(* Logix 5000 project; controller PLC_MCC1300_75F1 vendor 1 type 14 code 166 rev 32.11; software revision 32.04; part 27 of 83 *)
(* tags used below, declared in another part *)
   GP_OB_InitializeMain : GP_OB_Initialize;
   M302SpeedUp : MAC_SpeedUp;
   M351 : MAC_Conveyor;
   M352 : MAC_Conveyor;
   M352_ALM : MAC_Conveyor_ALM;
   M352_Data : UDT_Convoy_SL;
   M352_HMR : MAC_Conveyor_HMR;
   M352_HMW : MAC_Conveyor_HMW;
   M352_INPUT_xSLFanOn : BOOL;
   M352_M1_DR : AXIS_CIP_DRIVE;
   M352_M1_DR_IN_MAJ : MOTION_INSTRUCTION;
   M352_M1_DR_IN_MAR : MOTION_INSTRUCTION;
   M352_M1_DR_IN_MAS : MOTION_INSTRUCTION;
   M352_M1_DR_IN_MRP : MOTION_INSTRUCTION;
   M352_M1_DR_MAFR : MOTION_INSTRUCTION;
   M352_M1_DR_MDR : MOTION_INSTRUCTION;
   M352_M1_DR_MSF : MOTION_INSTRUCTION;
   M352_M1_DR_MSO : MOTION_INSTRUCTION;
   M352_M1_DR_OUT_MAJ : MOTION_INSTRUCTION;
   M352_M1_DR_OUT_MAM : MOTION_INSTRUCTION;
   M352_M1_DR_OUT_MAR : MOTION_INSTRUCTION;
   M352_M1_DR_OUT_MAS : MOTION_INSTRUCTION;
   M352_M1_DR_OUT_MCD : MOTION_INSTRUCTION;
   M352_M1_DR_OUT_MRP : MOTION_INSTRUCTION;
   M352_ONS1 : BOOL;
   M352_Output_xAutoMode : BOOL;
   M352_Output_xDescentBlockGlass : BOOL;
   M352_Output_xGlassPresence : BOOL;
   M352_Output_xHA_Alarm : BOOL;   // W254HA1. Acustic alarm
   M352_Output_xHL_Alarm : BOOL;
   M352_Output_xRiseBlockGlass : BOOL;
   M352_SpaceConv_Utilities : SpaceConv_Utilities;
   TMP_d : DINT;
   TMP_dDirection : DINT;
   TMP_r : REAL;
   TMP_rAcc : REAL;
   TMP_rDec : REAL;
   TMP_rSpeed : REAL;
   TMP_rTarget_M1 : REAL;
   TMP_xForwardCommadnForCleaningZone : BOOL;
   TMP_xPositioning : BOOL;
   TMP_xPositioning_M1 : BOOL;
   TMP_xPowerSaving : BOOL;
   TMP_xReverse : BOOL;
   TMP_xReverse_M1 : BOOL;
   TMP_xRun : BOOL;
   TMP_xRun_M1 : BOOL;
   xAlwaysOFF : BOOL;
   Z300_Conveyor : UDT_StandConv[29];
   Z300_Conveyor_Conf : UDT_Conveyor_Config[29];
   Z300_Conveyor_HMW : MAC_Conveyor_ZC_HMW[29];
   Z300_Conveyor_IN_MOTION : MAC_Conveyor_ZC_IN_MOTION[29];
   Z301_HMR : MAC_Zone_ML_HMR;
   Z900 : MAC_Zone;
   Z900_HMW : MAC_Zone_HMW;
(* CommandLogic, continued *)

ROUTINE M352_Output   (* ladder *)
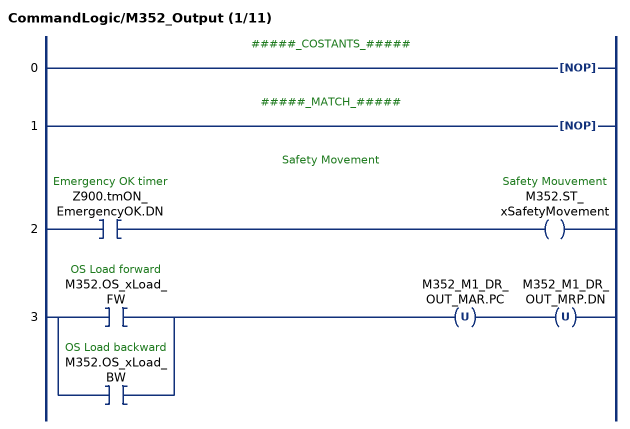
   // #####_COSTANTS_#####
   0: NOP();
   // #####_MATCH_#####
   1: NOP();
   // Safety Movement
   2: XIC(Z900.tmON_EmergencyOK.DN)OTE(M352.ST_xSafetyMovement);
   3: [XIC(M352.OS_xLoad_FW) ,XIC(M352.OS_xLoad_BW) ]OTU(M352_M1_DR_OUT_MAR.PC)OTU(M352_M1_DR_OUT_MRP.DN);
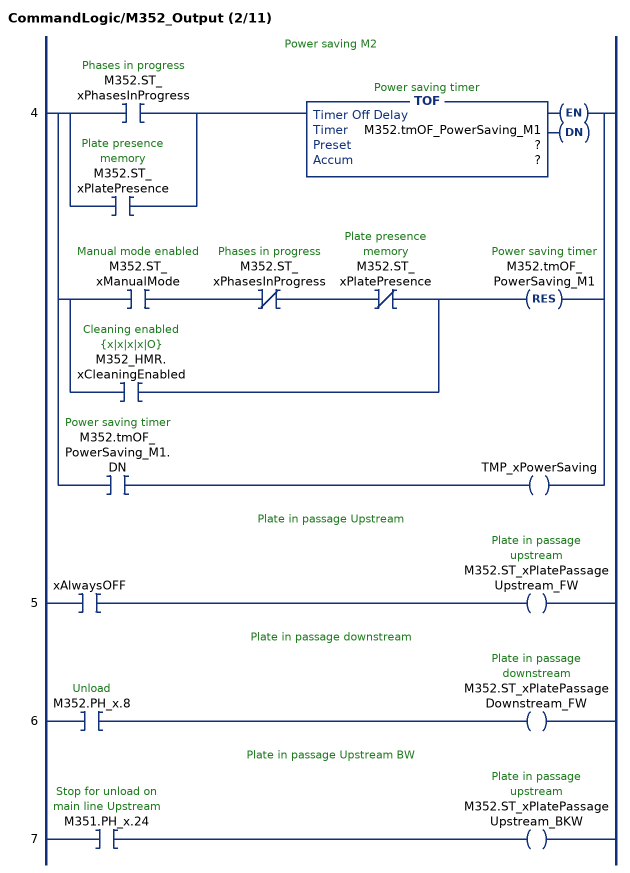
   // Power saving M2
   4: [[XIC(M352.ST_xPhasesInProgress) ,XIC(M352.ST_xPlatePresence) ] TOF(M352.tmOF_PowerSaving_M1,?,?) ,[XIC(M352.ST_xManualMode) XIO(M352.ST_xPhasesInProgress) XIO(M352.ST_xPlatePresence) ,XIC(M352_HMR.xCleaningEnabled) ] RES(M352.tmOF_PowerSaving_M1) ,XIC(M352.tmOF_PowerSaving_M1.DN) OTE(TMP_xPowerSaving) ];
   // Plate in passage Upstream
   5: XIC(xAlwaysOFF)OTE(M352.ST_xPlatePassageUpstream_FW);
   // Plate in passage downstream
   6: XIC(M352.PH_x.8)OTE(M352.ST_xPlatePassageDownstream_FW);
   // Plate in passage Upstream BW
   7: XIC(M351.PH_x.24)OTE(M352.ST_xPlatePassageUpstream_BKW);
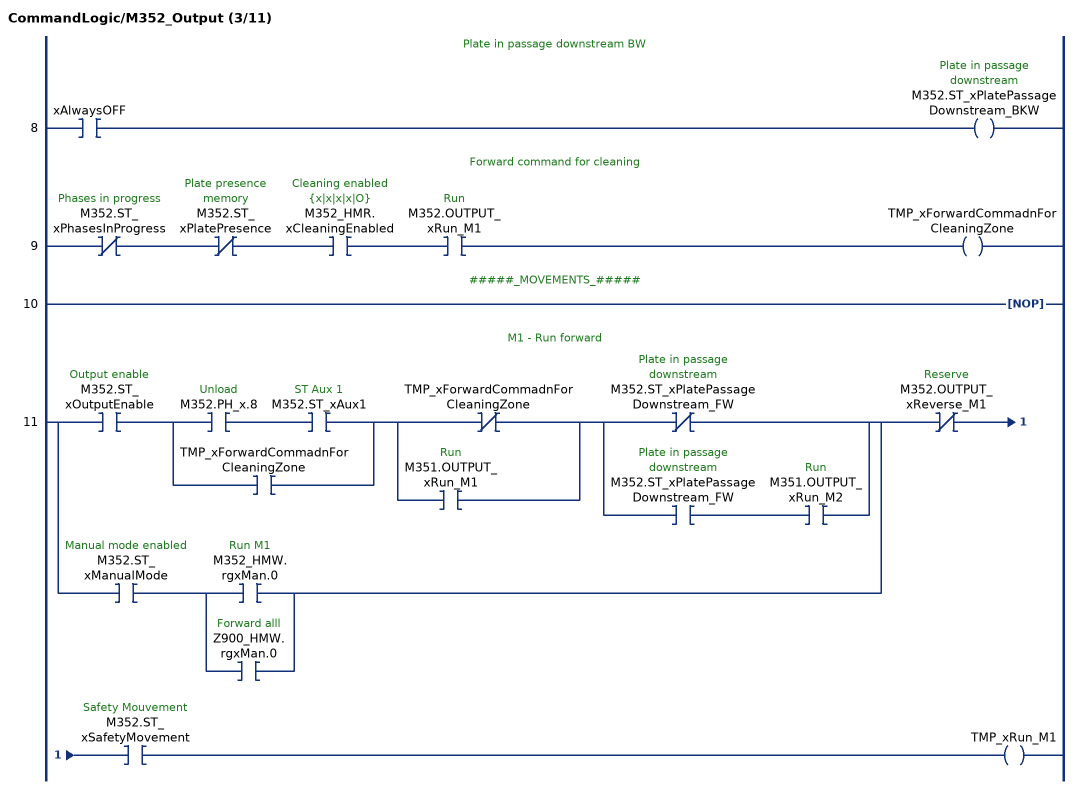
   // Plate in passage downstream BW
   8: XIC(xAlwaysOFF)OTE(M352.ST_xPlatePassageDownstream_BKW);
   // Forward command for cleaning
   9: XIO(M352.ST_xPhasesInProgress)XIO(M352.ST_xPlatePresence)XIC(M352_HMR.xCleaningEnabled)XIC(M352.OUTPUT_xRun_M1)OTE(TMP_xForwardCommadnForCleaningZone);
   // #####_MOVEMENTS_#####
   10: NOP();
   // M1 - Run forward
   11: [XIC(M352.ST_xOutputEnable) [XIC(M352.PH_x.8) XIC(M352.ST_xAux1) ,XIC(TMP_xForwardCommadnForCleaningZone) ] [XIO(TMP_xForwardCommadnForCleaningZone) ,XIC(M351.OUTPUT_xRun_M1) ] [XIO(M352.ST_xPlatePassageDownstream_FW) ,XIC(M352.ST_xPlatePassageDownstream_FW) XIC(M351.OUTPUT_xRun_M2) ] ,XIC(M352.ST_xManualMode) [XIC(M352_HMW.rgxMan.0) ,XIC(Z900_HMW.rgxMan.0) ] ]XIO(M352.OUTPUT_xReverse_M1)XIC(M352.ST_xSafetyMovement)OTE(TMP_xRun_M1);
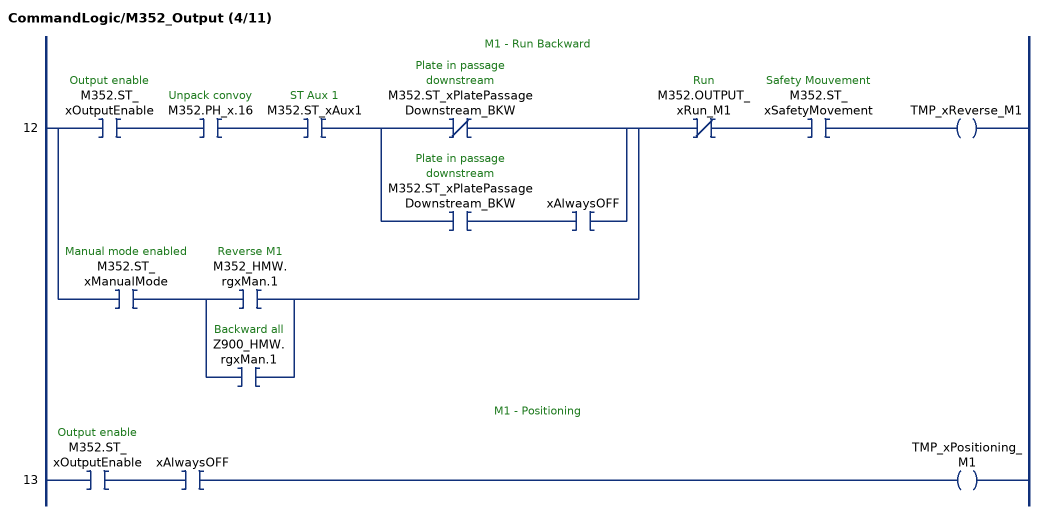
   // M1 - Run Backward
   12: [XIC(M352.ST_xOutputEnable) XIC(M352.PH_x.16) XIC(M352.ST_xAux1) [XIO(M352.ST_xPlatePassageDownstream_BKW) ,XIC(M352.ST_xPlatePassageDownstream_BKW) XIC(xAlwaysOFF) ] ,XIC(M352.ST_xManualMode) [XIC(M352_HMW.rgxMan.1) ,XIC(Z900_HMW.rgxMan.1) ] ]XIO(M352.OUTPUT_xRun_M1)XIC(M352.ST_xSafetyMovement)OTE(TMP_xReverse_M1);
   // M1 - Positioning
   13: XIC(M352.ST_xOutputEnable)XIC(xAlwaysOFF)OTE(TMP_xPositioning_M1);
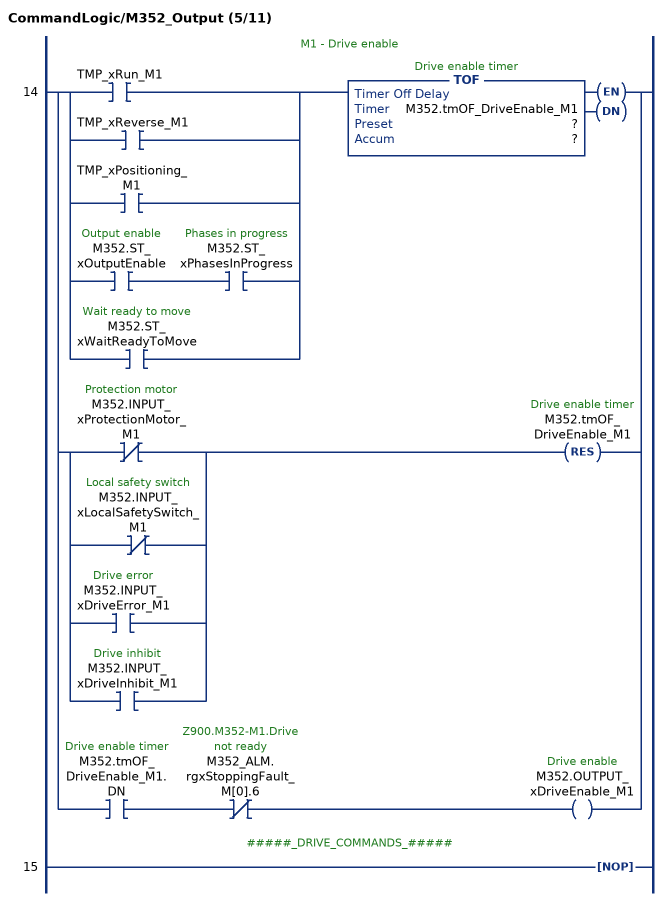
   // M1 - Drive enable
   14: [[XIC(TMP_xRun_M1) ,XIC(TMP_xReverse_M1) ,XIC(TMP_xPositioning_M1) ,XIC(M352.ST_xOutputEnable) XIC(M352.ST_xPhasesInProgress) ,XIC(M352.ST_xWaitReadyToMove) ] TOF(M352.tmOF_DriveEnable_M1,?,?) ,[XIO(M352.INPUT_xProtectionMotor_M1) ,XIO(M352.INPUT_xLocalSafetySwitch_M1) ,XIC(M352.INPUT_xDriveError_M1) ,XIC(M352.INPUT_xDriveInhibit_M1) ] RES(M352.tmOF_DriveEnable_M1) ,XIC(M352.tmOF_DriveEnable_M1.DN) XIO(M352_ALM.rgxStoppingFault_M[0].6) OTE(M352.OUTPUT_xDriveEnable_M1) ];
   // #####_DRIVE_COMMANDS_#####
   15: NOP();
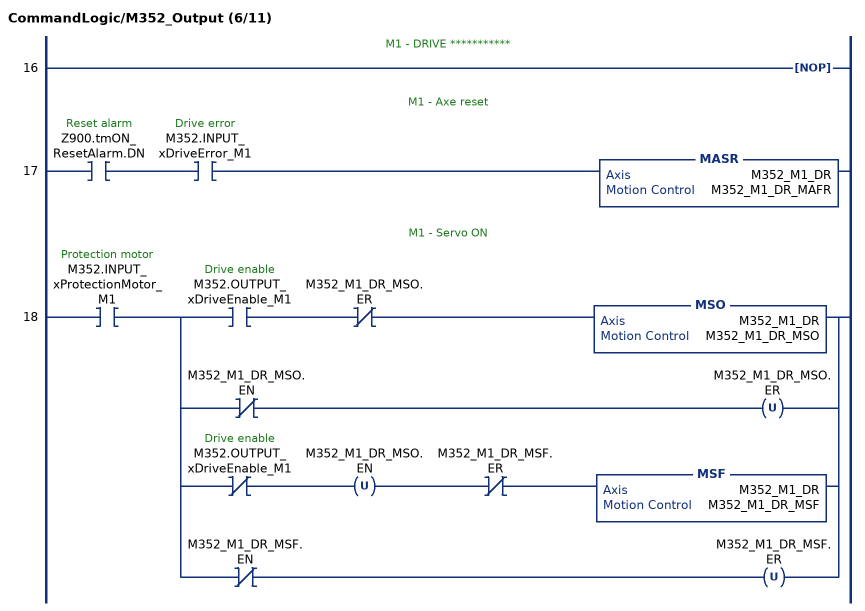
   // M1 - DRIVE ***********
   16: NOP();
   // M1 - Axe reset
   17: XIC(Z900.tmON_ResetAlarm.DN)XIC(M352.INPUT_xDriveError_M1)MASR(M352_M1_DR,M352_M1_DR_MAFR);
   // M1 - Servo ON
   18: XIC(M352.INPUT_xProtectionMotor_M1)[XIC(M352.OUTPUT_xDriveEnable_M1) XIO(M352_M1_DR_MSO.ER) MSO(M352_M1_DR,M352_M1_DR_MSO) ,XIO(M352_M1_DR_MSO.EN) OTU(M352_M1_DR_MSO.ER) ,XIO(M352.OUTPUT_xDriveEnable_M1) OTU(M352_M1_DR_MSO.EN) XIO(M352_M1_DR_MSF.ER) MSF(M352_M1_DR,M352_M1_DR_MSF) ,XIO(M352_M1_DR_MSF.EN) OTU(M352_M1_DR_MSF.ER) ];
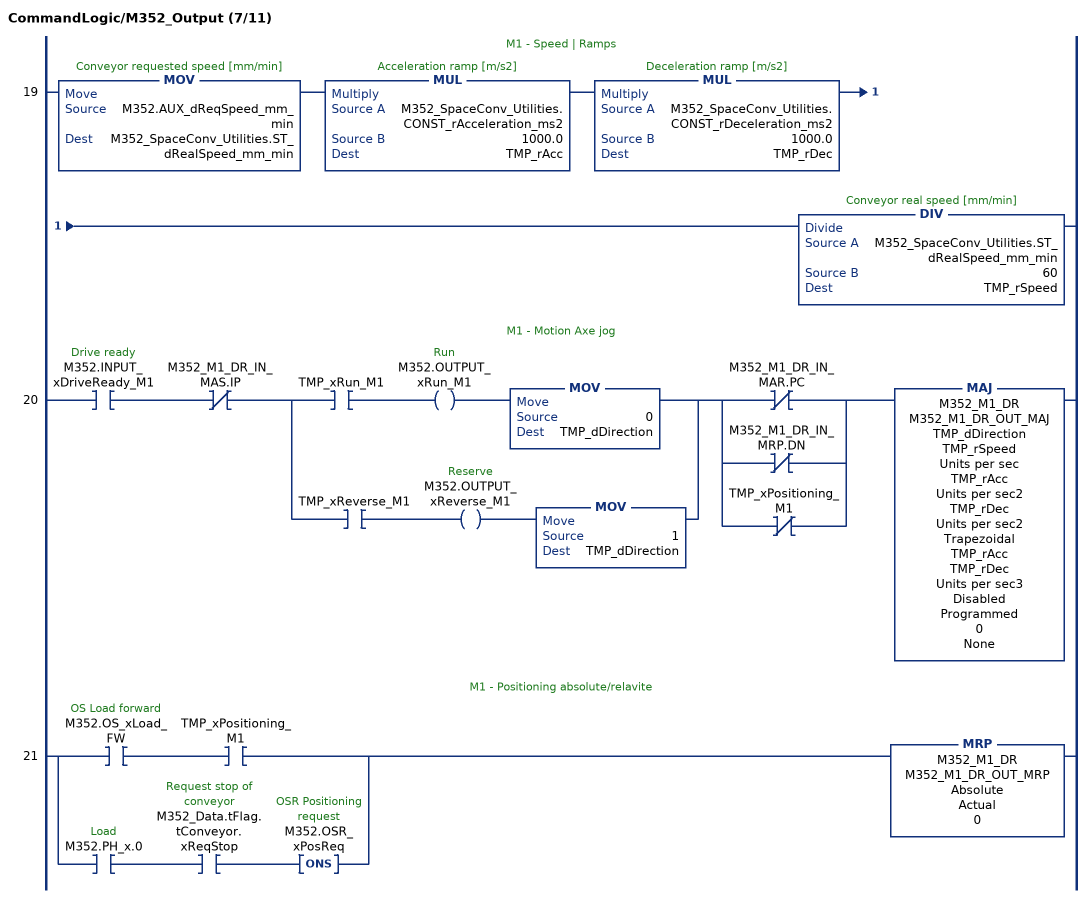
   // M1 - Speed | Ramps
   19: MOV(M352.AUX_dReqSpeed_mm_min,M352_SpaceConv_Utilities.ST_dRealSpeed_mm_min)MUL(M352_SpaceConv_Utilities.CONST_rAcceleration_ms2,1000.0,TMP_rAcc)MUL(M352_SpaceConv_Utilities.CONST_rDeceleration_ms2,1000.0,TMP_rDec)DIV(M352_SpaceConv_Utilities.ST_dRealSpeed_mm_min,60,TMP_rSpeed);
   // M1 - Motion Axe jog
   20: XIC(M352.INPUT_xDriveReady_M1)XIO(M352_M1_DR_IN_MAS.IP)[XIC(TMP_xRun_M1) OTE(M352.OUTPUT_xRun_M1) MOV(0,TMP_dDirection) ,XIC(TMP_xReverse_M1) OTE(M352.OUTPUT_xReverse_M1) MOV(1,TMP_dDirection) ][XIO(M352_M1_DR_IN_MAR.PC) ,XIO(M352_M1_DR_IN_MRP.DN) ,XIO(TMP_xPositioning_M1) ]MAJ(M352_M1_DR,M352_M1_DR_OUT_MAJ,TMP_dDirection,TMP_rSpeed,Units per sec,TMP_rAcc,Units per sec2,TMP_rDec,Units per sec2,Trapezoidal,TMP_rAcc,TMP_rDec,Units per sec3,Disabled,Programmed,0,None);
   // M1 - Positioning absolute/relavite
   21: [XIC(M352.OS_xLoad_FW) XIC(TMP_xPositioning_M1) ,XIC(M352.PH_x.0) XIC(M352_Data.tFlag.tConveyor.xReqStop) ONS(M352.OSR_xPosReq) ]MRP(M352_M1_DR,M352_M1_DR_OUT_MRP,Absolute,Actual,0);
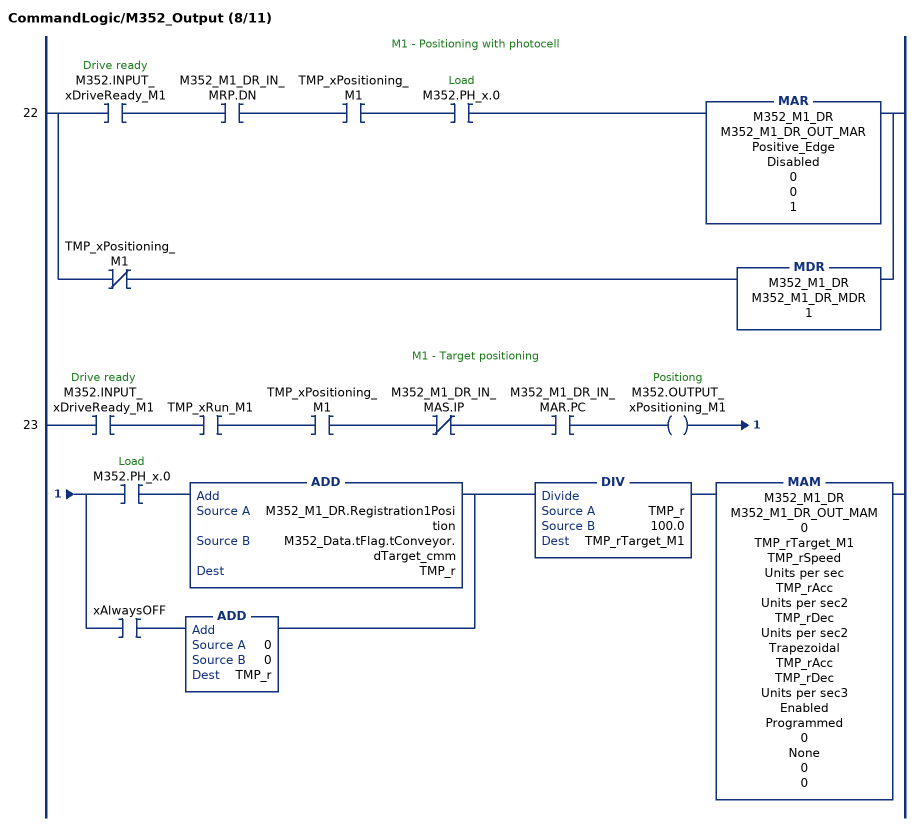
   // M1 - Positioning with photocell
   22: [XIC(M352.INPUT_xDriveReady_M1) XIC(M352_M1_DR_IN_MRP.DN) XIC(TMP_xPositioning_M1) XIC(M352.PH_x.0) MAR(M352_M1_DR,M352_M1_DR_OUT_MAR,Positive_Edge,Disabled,0,0,1) ,XIO(TMP_xPositioning_M1) MDR(M352_M1_DR,M352_M1_DR_MDR,1) ];
   // M1 - Target positioning
   23: XIC(M352.INPUT_xDriveReady_M1)XIC(TMP_xRun_M1)XIC(TMP_xPositioning_M1)XIO(M352_M1_DR_IN_MAS.IP)XIC(M352_M1_DR_IN_MAR.PC)OTE(M352.OUTPUT_xPositioning_M1)[XIC(M352.PH_x.0) ADD(M352_M1_DR.Registration1Position,M352_Data.tFlag.tConveyor.dTarget_cmm,TMP_r) ,XIC(xAlwaysOFF) ADD(0,0,TMP_r) ]DIV(TMP_r,100.0,TMP_rTarget_M1)MAM(M352_M1_DR,M352_M1_DR_OUT_MAM,0,TMP_rTarget_M1,TMP_rSpeed,Units per sec,TMP_rAcc,Units per sec2,TMP_rDec,Units per sec2,Trapezoidal,TMP_rAcc,TMP_rDec,Units per sec3,Enabled,Programmed,0,None,0,0);
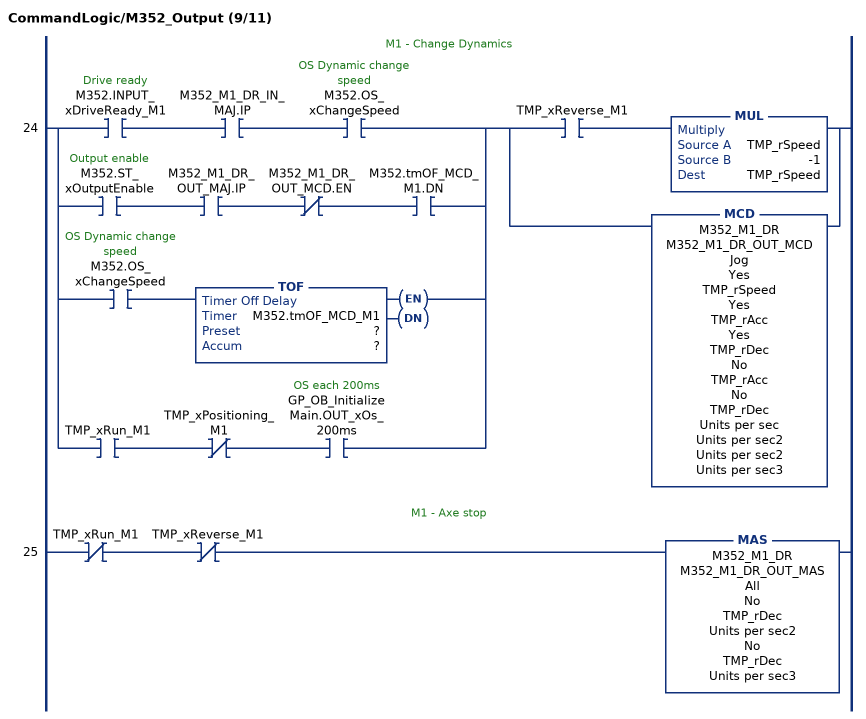
   // M1 - Change Dynamics
   24: [XIC(M352.INPUT_xDriveReady_M1) XIC(M352_M1_DR_IN_MAJ.IP) XIC(M352.OS_xChangeSpeed) ,XIC(M352.ST_xOutputEnable) XIC(M352_M1_DR_OUT_MAJ.IP) XIO(M352_M1_DR_OUT_MCD.EN) XIC(M352.tmOF_MCD_M1.DN) ,XIC(M352.OS_xChangeSpeed) TOF(M352.tmOF_MCD_M1,?,?) ,XIC(TMP_xRun_M1) XIO(TMP_xPositioning_M1) XIC(GP_OB_InitializeMain.OUT_xOs_200ms) ][XIC(TMP_xReverse_M1) MUL(TMP_rSpeed,-1,TMP_rSpeed) ,MCD(M352_M1_DR,M352_M1_DR_OUT_MCD,Jog,Yes,TMP_rSpeed,Yes,TMP_rAcc,Yes,TMP_rDec,No,TMP_rAcc,No,TMP_rDec,Units per sec,Units per sec2,Units per sec2,Units per sec3) ];
   // M1 - Axe stop
   25: XIO(TMP_xRun_M1)XIO(TMP_xReverse_M1)MAS(M352_M1_DR,M352_M1_DR_OUT_MAS,All,No,TMP_rDec,Units per sec2,No,TMP_rDec,Units per sec3);
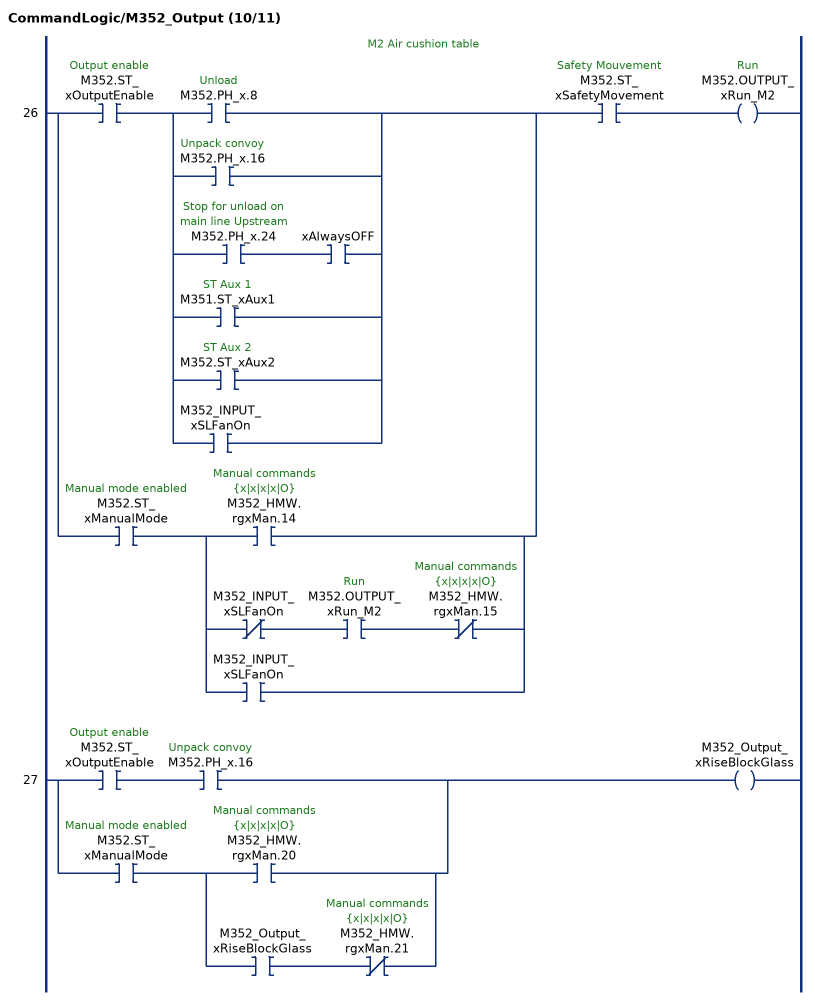
   // M2 Air cushion table
   26: [XIC(M352.ST_xOutputEnable) [XIC(M352.PH_x.8) ,XIC(M352.PH_x.16) ,XIC(M352.PH_x.24) XIC(xAlwaysOFF) ,XIC(M351.ST_xAux1) ,XIC(M352.ST_xAux2) ,XIC(M352_INPUT_xSLFanOn) ] ,XIC(M352.ST_xManualMode) [XIC(M352_HMW.rgxMan.14) ,XIO(M352_INPUT_xSLFanOn) XIC(M352.OUTPUT_xRun_M2) XIO(M352_HMW.rgxMan.15) ,XIC(M352_INPUT_xSLFanOn) ] ]XIC(M352.ST_xSafetyMovement)OTE(M352.OUTPUT_xRun_M2);
   27: [XIC(M352.ST_xOutputEnable) XIC(M352.PH_x.16) ,XIC(M352.ST_xManualMode) [XIC(M352_HMW.rgxMan.20) ,XIC(M352_Output_xRiseBlockGlass) XIO(M352_HMW.rgxMan.21) ] ]OTE(M352_Output_xRiseBlockGlass);
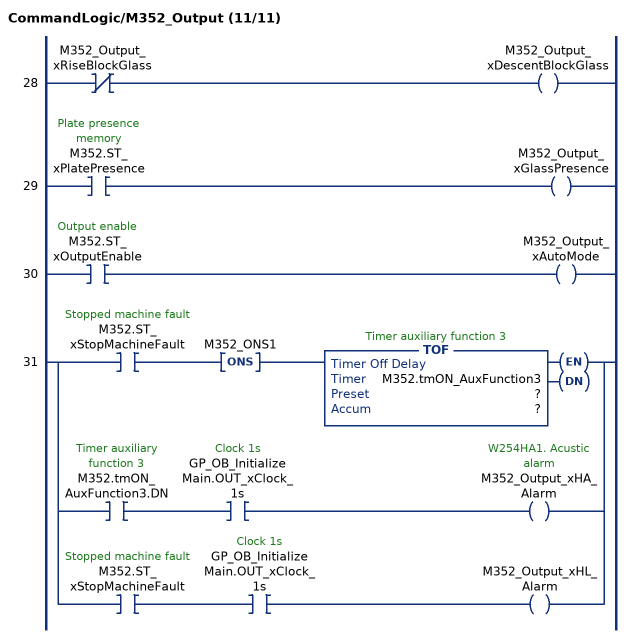
   28: XIO(M352_Output_xRiseBlockGlass)OTE(M352_Output_xDescentBlockGlass);
   29: XIC(M352.ST_xPlatePresence)OTE(M352_Output_xGlassPresence);
   30: XIC(M352.ST_xOutputEnable)OTE(M352_Output_xAutoMode);
   31: [XIC(M352.ST_xStopMachineFault) ONS(M352_ONS1) TOF(M352.tmON_AuxFunction3,?,?) ,XIC(M352.tmON_AuxFunction3.DN) XIC(GP_OB_InitializeMain.OUT_xClock_1s) OTE(M352_Output_xHA_Alarm) ,XIC(M352.ST_xStopMachineFault) XIC(GP_OB_InitializeMain.OUT_xClock_1s) OTE(M352_Output_xHL_Alarm) ];
END_ROUTINE

ROUTINE M360M1_Conveyor_Output   (* ladder *)
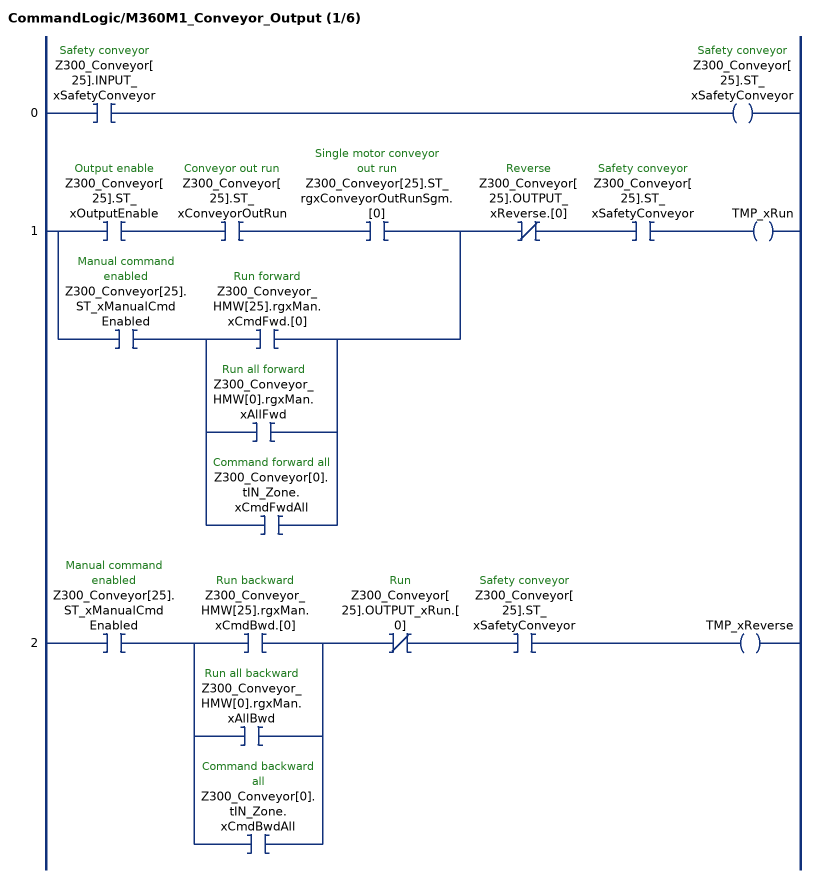
   0: XIC(Z300_Conveyor[25].INPUT_xSafetyConveyor)OTE(Z300_Conveyor[25].ST_xSafetyConveyor);
   1: [XIC(Z300_Conveyor[25].ST_xOutputEnable) XIC(Z300_Conveyor[25].ST_xConveyorOutRun) XIC(Z300_Conveyor[25].ST_rgxConveyorOutRunSgm.[0]) ,XIC(Z300_Conveyor[25].ST_xManualCmdEnabled) [XIC(Z300_Conveyor_HMW[25].rgxMan.xCmdFwd.[0]) ,XIC(Z300_Conveyor_HMW[0].rgxMan.xAllFwd) ,XIC(Z300_Conveyor[0].tIN_Zone.xCmdFwdAll) ] ]XIO(Z300_Conveyor[25].OUTPUT_xReverse.[0])XIC(Z300_Conveyor[25].ST_xSafetyConveyor)OTE(TMP_xRun);
   2: XIC(Z300_Conveyor[25].ST_xManualCmdEnabled)[XIC(Z300_Conveyor_HMW[25].rgxMan.xCmdBwd.[0]) ,XIC(Z300_Conveyor_HMW[0].rgxMan.xAllBwd) ,XIC(Z300_Conveyor[0].tIN_Zone.xCmdBwdAll) ]XIO(Z300_Conveyor[25].OUTPUT_xRun.[0])XIC(Z300_Conveyor[25].ST_xSafetyConveyor)OTE(TMP_xReverse);
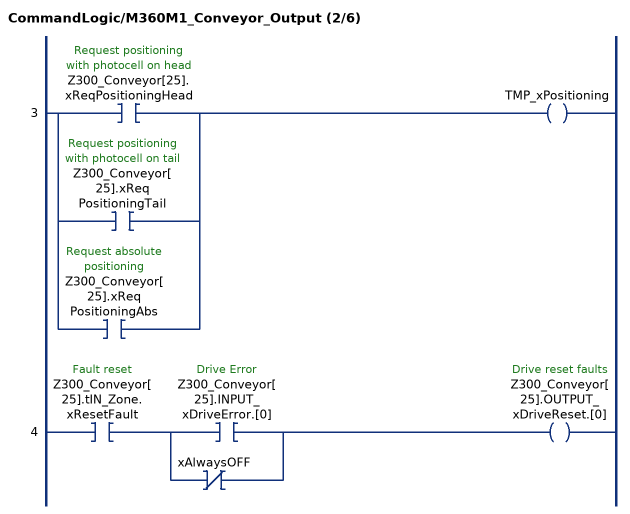
   3: [XIC(Z300_Conveyor[25].xReqPositioningHead) ,XIC(Z300_Conveyor[25].xReqPositioningTail) ,XIC(Z300_Conveyor[25].xReqPositioningAbs) ]OTE(TMP_xPositioning);
   4: XIC(Z300_Conveyor[25].tIN_Zone.xResetFault)[XIC(Z300_Conveyor[25].INPUT_xDriveError.[0]) ,XIO(xAlwaysOFF) ]OTE(Z300_Conveyor[25].OUTPUT_xDriveReset.[0]);
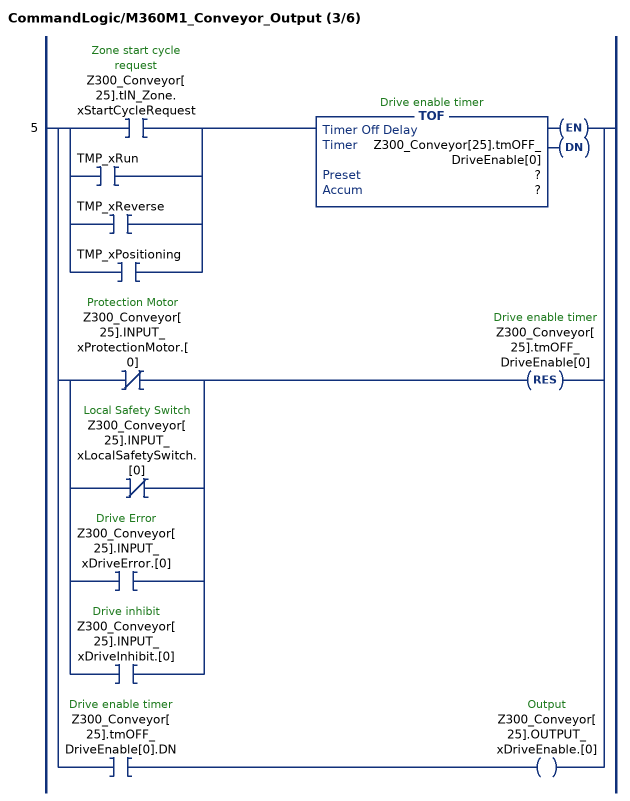
   5: [[XIC(Z300_Conveyor[25].tIN_Zone.xStartCycleRequest) ,XIC(TMP_xRun) ,XIC(TMP_xReverse) ,XIC(TMP_xPositioning) ] TOF(Z300_Conveyor[25].tmOFF_DriveEnable[0],?,?) ,[XIO(Z300_Conveyor[25].INPUT_xProtectionMotor.[0]) ,XIO(Z300_Conveyor[25].INPUT_xLocalSafetySwitch.[0]) ,XIC(Z300_Conveyor[25].INPUT_xDriveError.[0]) ,XIC(Z300_Conveyor[25].INPUT_xDriveInhibit.[0]) ] RES(Z300_Conveyor[25].tmOFF_DriveEnable[0]) ,XIC(Z300_Conveyor[25].tmOFF_DriveEnable[0].DN) OTE(Z300_Conveyor[25].OUTPUT_xDriveEnable.[0]) ];
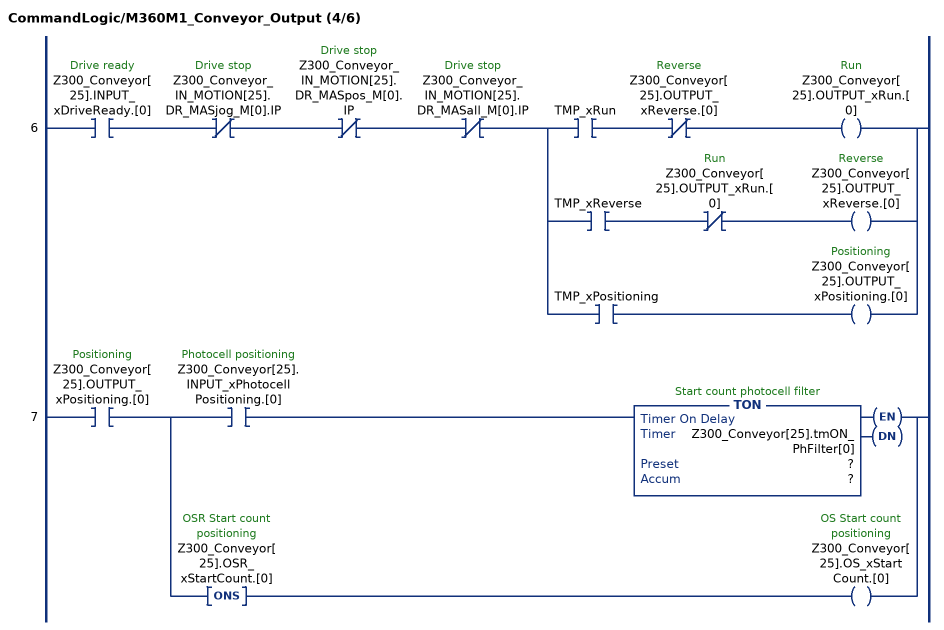
   6: XIC(Z300_Conveyor[25].INPUT_xDriveReady.[0])XIO(Z300_Conveyor_IN_MOTION[25].DR_MASjog_M[0].IP)XIO(Z300_Conveyor_IN_MOTION[25].DR_MASpos_M[0].IP)XIO(Z300_Conveyor_IN_MOTION[25].DR_MASall_M[0].IP)[XIC(TMP_xRun) XIO(Z300_Conveyor[25].OUTPUT_xReverse.[0]) OTE(Z300_Conveyor[25].OUTPUT_xRun.[0]) ,XIC(TMP_xReverse) XIO(Z300_Conveyor[25].OUTPUT_xRun.[0]) OTE(Z300_Conveyor[25].OUTPUT_xReverse.[0]) ,XIC(TMP_xPositioning) OTE(Z300_Conveyor[25].OUTPUT_xPositioning.[0]) ];
   7: XIC(Z300_Conveyor[25].OUTPUT_xPositioning.[0])[XIC(Z300_Conveyor[25].INPUT_xPhotocellPositioning.[0]) TON(Z300_Conveyor[25].tmON_PhFilter[0],?,?) ,ONS(Z300_Conveyor[25].OSR_xStartCount.[0]) OTE(Z300_Conveyor[25].OS_xStartCount.[0]) ];
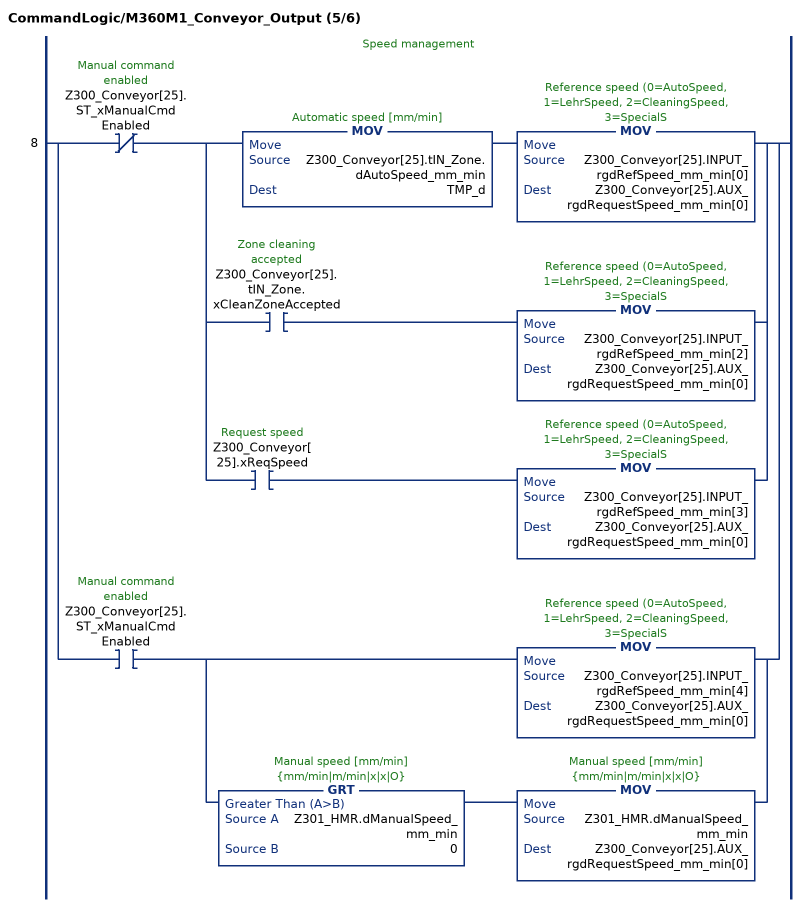
   // Speed management
   8: [XIO(Z300_Conveyor[25].ST_xManualCmdEnabled) [MOV(Z300_Conveyor[25].tIN_Zone.dAutoSpeed_mm_min,TMP_d) MOV(Z300_Conveyor[25].INPUT_rgdRefSpeed_mm_min[0],Z300_Conveyor[25].AUX_rgdRequestSpeed_mm_min[0]) ,XIC(Z300_Conveyor[25].tIN_Zone.xCleanZoneAccepted) MOV(Z300_Conveyor[25].INPUT_rgdRefSpeed_mm_min[2],Z300_Conveyor[25].AUX_rgdRequestSpeed_mm_min[0]) ,XIC(Z300_Conveyor[25].xReqSpeed) MOV(Z300_Conveyor[25].INPUT_rgdRefSpeed_mm_min[3],Z300_Conveyor[25].AUX_rgdRequestSpeed_mm_min[0]) ] ,XIC(Z300_Conveyor[25].ST_xManualCmdEnabled) [MOV(Z300_Conveyor[25].INPUT_rgdRefSpeed_mm_min[4],Z300_Conveyor[25].AUX_rgdRequestSpeed_mm_min[0]) ,GRT(Z301_HMR.dManualSpeed_mm_min,0) MOV(Z301_HMR.dManualSpeed_mm_min,Z300_Conveyor[25].AUX_rgdRequestSpeed_mm_min[0]) ] ];
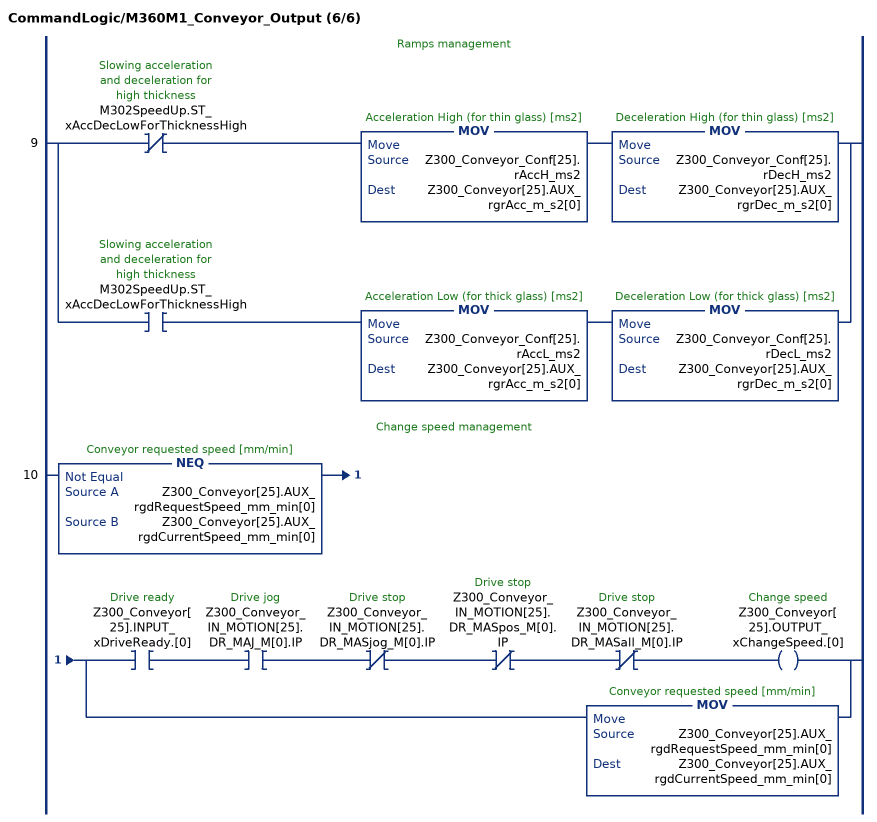
   // Ramps management
   9: [XIO(M302SpeedUp.ST_xAccDecLowForThicknessHigh) MOV(Z300_Conveyor_Conf[25].rAccH_ms2,Z300_Conveyor[25].AUX_rgrAcc_m_s2[0]) MOV(Z300_Conveyor_Conf[25].rDecH_ms2,Z300_Conveyor[25].AUX_rgrDec_m_s2[0]) ,XIC(M302SpeedUp.ST_xAccDecLowForThicknessHigh) MOV(Z300_Conveyor_Conf[25].rAccL_ms2,Z300_Conveyor[25].AUX_rgrAcc_m_s2[0]) MOV(Z300_Conveyor_Conf[25].rDecL_ms2,Z300_Conveyor[25].AUX_rgrDec_m_s2[0]) ];
   // Change speed management
   10: NEQ(Z300_Conveyor[25].AUX_rgdRequestSpeed_mm_min[0],Z300_Conveyor[25].AUX_rgdCurrentSpeed_mm_min[0])[XIC(Z300_Conveyor[25].INPUT_xDriveReady.[0]) XIC(Z300_Conveyor_IN_MOTION[25].DR_MAJ_M[0].IP) XIO(Z300_Conveyor_IN_MOTION[25].DR_MASjog_M[0].IP) XIO(Z300_Conveyor_IN_MOTION[25].DR_MASpos_M[0].IP) XIO(Z300_Conveyor_IN_MOTION[25].DR_MASall_M[0].IP) OTE(Z300_Conveyor[25].OUTPUT_xChangeSpeed.[0]) ,MOV(Z300_Conveyor[25].AUX_rgdRequestSpeed_mm_min[0],Z300_Conveyor[25].AUX_rgdCurrentSpeed_mm_min[0]) ];
END_ROUTINE

ROUTINE Main   (* ladder *)
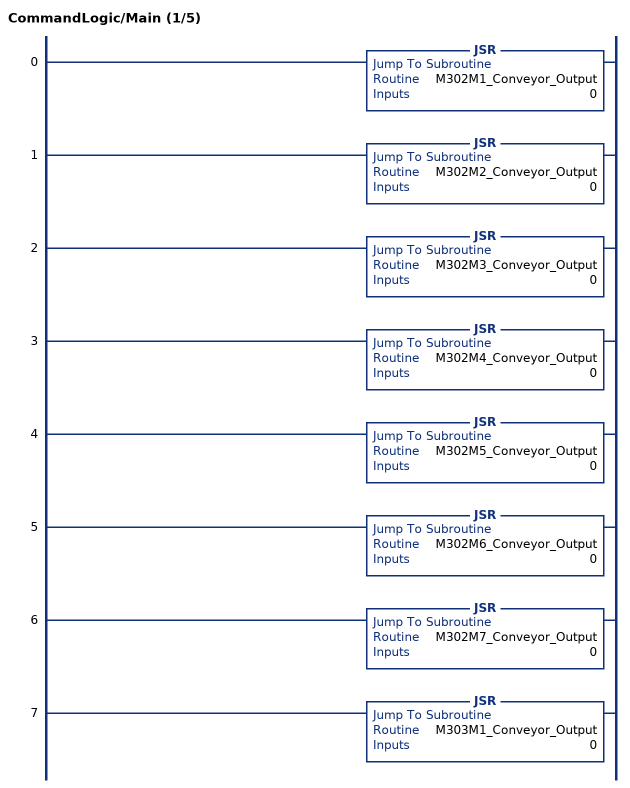
   0: JSR(M302M1_Conveyor_Output,0);
   1: JSR(M302M2_Conveyor_Output,0);
   2: JSR(M302M3_Conveyor_Output,0);
   3: JSR(M302M4_Conveyor_Output,0);
   4: JSR(M302M5_Conveyor_Output,0);
   5: JSR(M302M6_Conveyor_Output,0);
   6: JSR(M302M7_Conveyor_Output,0);
   7: JSR(M303M1_Conveyor_Output,0);
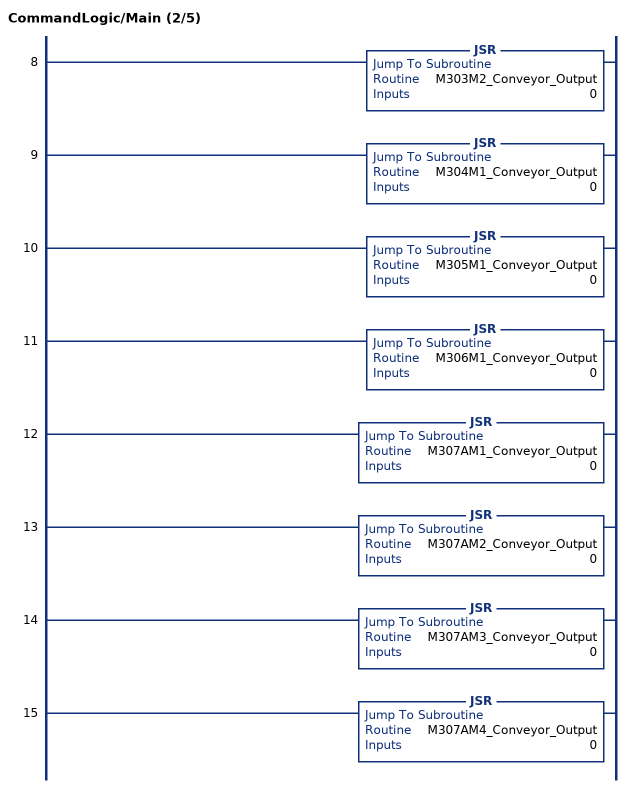
   8: JSR(M303M2_Conveyor_Output,0);
   9: JSR(M304M1_Conveyor_Output,0);
   10: JSR(M305M1_Conveyor_Output,0);
   11: JSR(M306M1_Conveyor_Output,0);
   12: JSR(M307AM1_Conveyor_Output,0);
   13: JSR(M307AM2_Conveyor_Output,0);
   14: JSR(M307AM3_Conveyor_Output,0);
   15: JSR(M307AM4_Conveyor_Output,0);
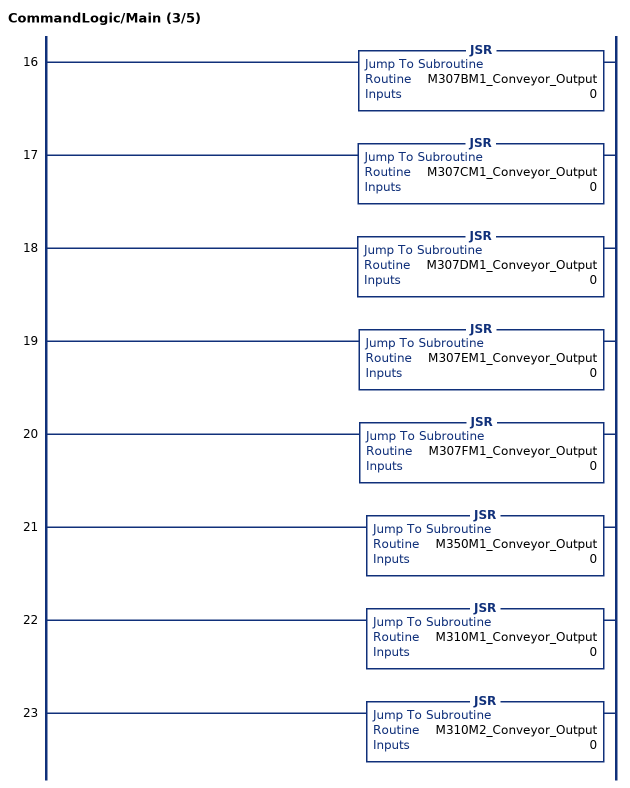
   16: JSR(M307BM1_Conveyor_Output,0);
   17: JSR(M307CM1_Conveyor_Output,0);
   18: JSR(M307DM1_Conveyor_Output,0);
   19: JSR(M307EM1_Conveyor_Output,0);
   20: JSR(M307FM1_Conveyor_Output,0);
   21: JSR(M350M1_Conveyor_Output,0);
   22: JSR(M310M1_Conveyor_Output,0);
   23: JSR(M310M2_Conveyor_Output,0);
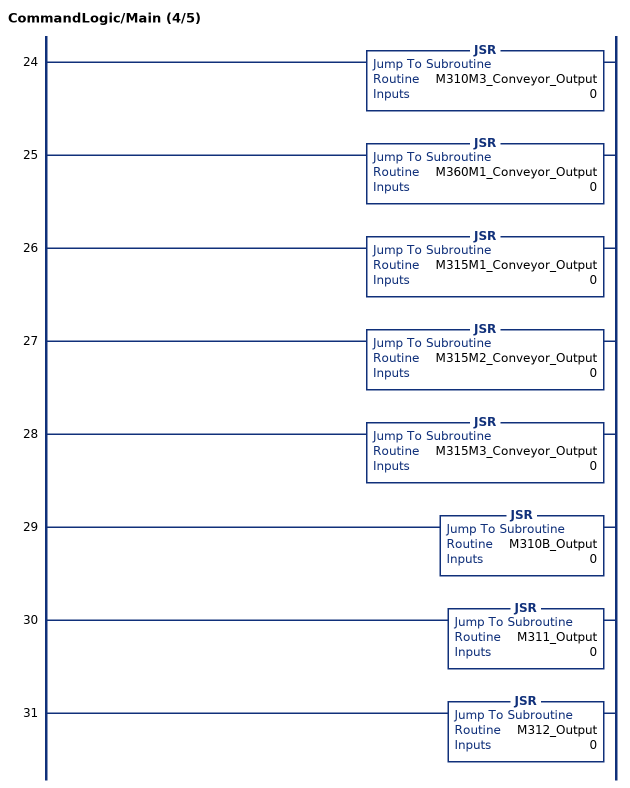
   24: JSR(M310M3_Conveyor_Output,0);
   25: JSR(M360M1_Conveyor_Output,0);
   26: JSR(M315M1_Conveyor_Output,0);
   27: JSR(M315M2_Conveyor_Output,0);
   28: JSR(M315M3_Conveyor_Output,0);
   29: JSR(M310B_Output,0);
   30: JSR(M311_Output,0);
   31: JSR(M312_Output,0);
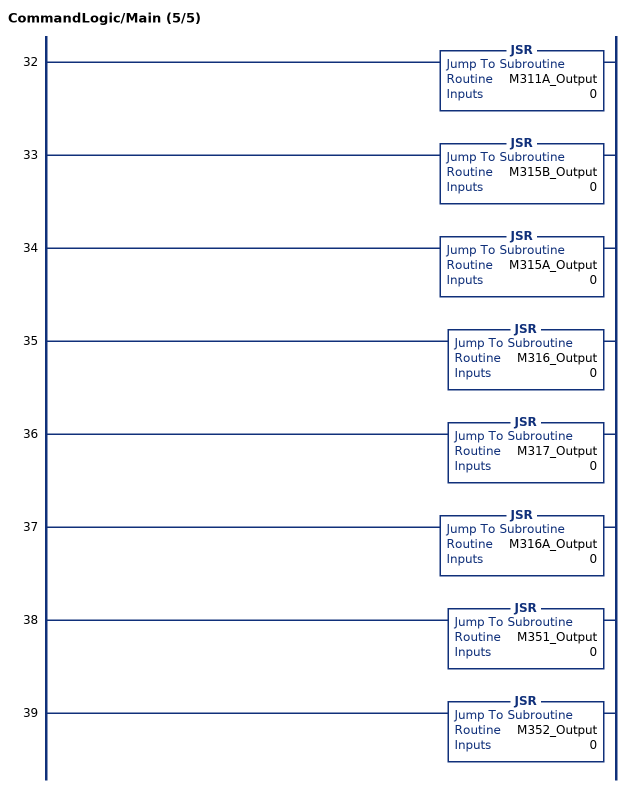
   32: JSR(M311A_Output,0);
   33: JSR(M315B_Output,0);
   34: JSR(M315A_Output,0);
   35: JSR(M316_Output,0);
   36: JSR(M317_Output,0);
   37: JSR(M316A_Output,0);
   38: JSR(M351_Output,0);
   39: JSR(M352_Output,0);
END_ROUTINE
END_PROGRAM
